(* Logix 5000 project; controller PLC_MCC1300_75F1 vendor 1 type 14 code 166 rev 32.11; software revision 32.04; part 5 of 83 *)
(* tags used below, declared in another part *)
   GP_PlateYPosition : GP_PlateYPosition;
   GP_PosWindow : GP_PosWindow;
   GP_RampManagement : GP_RampManagement;
   GP_RampSpace : GP_RampSpace;
   GP_ScadaPlate : GP_ScadaPlate;
   Gp_SpaceConvUtilities_V1 : GP_SpaceConvUtilities_V1;
   GP_TrackingAddCap : GP_TrackingAddCap;
   GP_TrackingFiring : GP_TrackingFiring;
   GP_TrackingFiringForConvoy : GP_TrackingFiringForConvoy;
   GP_TrackingGetFirstPlateInConveyor : GP_TrackingGetFirstPlateInConveyor;

ADD_ON_INSTRUCTION GP_PlateYPosition   (* revision 1.0 *)
VAR_IN_OUT
   INO_tPlateData : UDT_ConvoyCap_ZC; {required}
END_VAR
VAR_INPUT
   IN_dRequestGapLite_cmm : DINT; {access None, required}   // Requested gap between lites
   IN_dOffset_cmm : DINT; {access None, required}   // Position offset
   IN_xWander : BOOL; {access None, required}   // Calculate wander & total width
   IN_xBarycenter : BOOL; {access None, required}   // Calculate Barycenter
   IN_rgxNoGapLite : DINT; {access None, required}   // Consider gap of single lite [0:ConsiderGap, 1:NotConsiderGap]
END_VAR
VAR
   TMP_dLite : DINT; {access None}
   TMP_dMaxLites : DINT; {access None}
   TMP_dCapEdge_cmm : DINT; {access None}
END_VAR

ROUTINE Logic   (* structured text *)
   
   SIZE(INO_tPlateData.rgtCap[0].rgtLite[0],0,TMP_dMaxLites);
   IF INO_tPlateData.rgtCap[0].dID <> 0 THEN
       IF INO_tPlateData.rgtCap[0].dNumLites > 0 AND IN_xBarycenter THEN
           TMP_dCapEdge_cmm := (IN_dOffset_cmm + INO_tPlateData.rgtCap[0].dCutWander_cmm) - (INO_tPlateData.rgtCap[0].dWidth_cmm / 2) - (IN_dRequestGapLite_cmm / 2);
           FOR TMP_dLite := 0 TO TMP_dMaxLites - 1 DO
               IF INO_tPlateData.rgtCap[0].rgtLite[TMP_dLite].dID <> 0 THEN
                   INO_tPlateData.rgtCap[0].rgtLite[TMP_dLite].dBarycenter_cmm := TMP_dCapEdge_cmm + (INO_tPlateData.rgtCap[0].rgtLite[TMP_dLite].dWidth_cmm / 2);
                   IF NOT (IN_rgxNoGapLite.[TMP_dLite]) THEN
                       TMP_dCapEdge_cmm := TMP_dCapEdge_cmm + INO_tPlateData.rgtCap[0].rgtLite[TMP_dLite].dWidth_cmm + IN_dRequestGapLite_cmm;
   					//Update gap in cap data
   					INO_tPlateData.rgtCap[0].dGap_cmm := IN_dRequestGapLite_cmm;
                   ELSE
                       TMP_dCapEdge_cmm := TMP_dCapEdge_cmm + INO_tPlateData.rgtCap[0].rgtLite[TMP_dLite].dWidth_cmm;
                   END_IF;
               END_IF;
           END_FOR;
       ELSIF INO_tPlateData.rgtCap[0].dNumLites > 0 AND IN_xWander THEN
           FOR TMP_dLite := 0 TO TMP_dMaxLites - 1 DO
               IF INO_tPlateData.rgtCap[0].rgtLite[TMP_dLite].dID <> 0 THEN
                   TMP_dCapEdge_cmm := INO_tPlateData.rgtCap[0].rgtLite[TMP_dLite].dBarycenter_cmm - (INO_tPlateData.rgtCap[0].rgtLite[TMP_dLite].dWidth_cmm / 2);
               END_IF;
           END_FOR;
           FOR TMP_dLite := 0 TO TMP_dMaxLites - 1 DO
               IF INO_tPlateData.rgtCap[0].rgtLite[TMP_dLite].dID <> 0 THEN
                   INO_tPlateData.rgtCap[0].dWidth_cmm := (INO_tPlateData.rgtCap[0].rgtLite[TMP_dLite].dBarycenter_cmm + (INO_tPlateData.rgtCap[0].rgtLite[TMP_dLite].dWidth_cmm / 2)) - TMP_dCapEdge_cmm;
               END_IF;
           END_FOR;
           INO_tPlateData.rgtCap[0].dCutWander_cmm := (TMP_dCapEdge_cmm + (INO_tPlateData.rgtCap[0].dWidth_cmm / 2)) - IN_dOffset_cmm;
       END_IF;
   END_IF;
   
END_ROUTINE
END_ADD_ON_INSTRUCTION

ADD_ON_INSTRUCTION GP_PosWindow   (* revision 1.0 *)
VAR_INPUT
   IN_dTarget : DINT; {access None, required}   // Request position [user unit]
   IN_dActual : DINT; {access None, required}   // Actual position [user unit]
   IN_dTollerance : DINT; {access None, required}   // Tollerance window [user unit]
   IN_dMode : DINT; {access None, required}   // Type mode (0=Included, 1=Greater/Included, 2=Less/Includedl, 3=Greater, 4=Less)
END_VAR
VAR_OUTPUT
   OUT_xPositionReached : BOOL; {access None, required}   // Position reached
END_VAR
VAR
   TMP_dMaxValue : DINT; {access None}
   TMP_dMinValue : DINT; {access None}
END_VAR

ROUTINE Logic   (* structured text *)
   TMP_dMinValue := IN_dTarget - IN_dTollerance ;
   TMP_dMaxValue := IN_dTarget + IN_dTollerance ;
   
   CASE IN_dMode OF
   
   0:	IF IN_dActual >= TMP_dMinValue AND IN_dActual <= TMP_dMaxValue THEN
   
   		OUT_xPositionReached := 1 ;
   
   	ELSE
   
   		OUT_xPositionReached := 0 ;
   
   	END_IF;
   
   1:	IF IN_dActual >= TMP_dMinValue THEN
   
   		OUT_xPositionReached := 1 ;
   
   	ELSE
   
   		OUT_xPositionReached := 0 ;
   
   	END_IF;
   
   2:	IF IN_dActual <= TMP_dMaxValue THEN
   
   		OUT_xPositionReached := 1 ;
   
   	ELSE
   
   		OUT_xPositionReached := 0 ;
   
   	END_IF;
   
   3:	IF IN_dActual > TMP_dMinValue THEN
   
   		OUT_xPositionReached := 1 ;
   
   	ELSE
   
   		OUT_xPositionReached := 0 ;
   
   	END_IF;
   
   4:	IF IN_dActual < TMP_dMaxValue THEN
   
   		OUT_xPositionReached := 1 ;
   
   	ELSE
   
   		OUT_xPositionReached := 0 ;
   
   	END_IF;
   
   END_CASE;
   
   EnableOut := 1 ;
END_ROUTINE
END_ADD_ON_INSTRUCTION

ADD_ON_INSTRUCTION GP_RampManagement   (* revision 1.0 *)
VAR_INPUT
   IN_xRun : BOOL; {access None, required}   // Run command
   IN_dSpeed_Setpoint : DINT; {access None, required}   // Setpoint speed [mm/min]
   IN_rAcc : REAL; {access None, required}   // Acceleration [m/s2]
   IN_rDec : REAL; {access None, required}   // Deceleration [m/s2]
   IN_rScan : REAL; {access None, required}   // Previous scan [ms]
END_VAR
VAR_IN_OUT
   INO_rPV_Speed : REAL; {required}   // Processed speed value [mm/min]
END_VAR
VAR_OUTPUT
   OUT_dStep_cmm : DINT; {access None, required}   // Incremental step for each scan cycle [mm/100]
   OUT_xRampInProgress : BOOL; {access None, required}   // Acceleration/Deceleration ramp in progress
   OUT_xAccInProgress : BOOL; {access None, required}   // Acceleration ramp in progress
   OUT_xDecInProgress : BOOL; {access None, required}   // Deceleration ramp in progress
END_VAR
VAR_IN_OUT
   INO_rReminderStep : REAL; {required}   // Reminder Step [mm/min]
END_VAR
VAR
   TMP_rDecLim : REAL; {access None}   // Deceleration limit [mm/min]
   TMP_rAccLim : REAL; {access None}   // Acceleration limit [mm/min]
   TMP_rDecStep : REAL; {access None}   // Deceleration step [mm/min]
   TMP_rAccStep : REAL; {access None}   // Acceleration step [mm/min]
   TMP_rSpeed_Setpoint : REAL; {access None}   // Setpoint speed [mm/min]
   TMP_rScan : REAL; {access None}   // Previous scan [ms]
   TMP_rStep : REAL; {access None}   // Actual Step with reminder [mm/min]
   TMP_rStepRound : REAL; {access None}   // Actual Step with reminder [mm/min]
END_VAR

ROUTINE Logic   (* structured text *)
   //Initialize
   OUT_dStep_cmm := 0;
   TMP_rSpeed_Setpoint := IN_dSpeed_Setpoint;
   TMP_rScan := IN_rScan;
   OUT_xRampInProgress := 0;
   OUT_xAccInProgress := 0;
   OUT_xDecInProgress := 0;
   
   //Check Speed, Acceleration and Deceleration Values > 0
   
   IF TMP_rSpeed_Setpoint > 0.0 AND IN_rAcc > 0.0 AND IN_rDec > 0.0 THEN
   
       // Acceleration
       IF IN_xRun AND TMP_rSpeed_Setpoint > INO_rPV_Speed THEN
           TMP_rAccStep := IN_rAcc * TMP_rScan * 60.0;
           INO_rPV_Speed := INO_rPV_Speed + TMP_rAccStep;
           TMP_rAccLim := TMP_rSpeed_Setpoint + TMP_rAccStep;
           OUT_xRampInProgress := 1;
           OUT_xAccInProgress := 1;
   
           IF IN_xRun AND INO_rPV_Speed > TMP_rSpeed_Setpoint AND INO_rPV_Speed < TMP_rAccLim THEN
               INO_rPV_Speed := TMP_rSpeed_Setpoint;
           END_IF;
   
           // Deceleration
   
       ELSIF (IN_xRun AND TMP_rSpeed_Setpoint < INO_rPV_Speed) OR (NOT (IN_xRun) AND INO_rPV_Speed > 0.0) THEN
           TMP_rDecStep := IN_rDec * TMP_rScan * 60.0;
           INO_rPV_Speed := INO_rPV_Speed - TMP_rDecStep;
           TMP_rDecLim := TMP_rSpeed_Setpoint - TMP_rDecStep;
           OUT_xRampInProgress := 1;
           OUT_xDecInProgress := 1;
   
           IF IN_xRun AND INO_rPV_Speed < TMP_rSpeed_Setpoint AND INO_rPV_Speed > TMP_rDecLim THEN
               INO_rPV_Speed := TMP_rSpeed_Setpoint;
           END_IF;
       END_IF;
   
       // Delete PV_Speed If < 0
   
       IF INO_rPV_Speed < 0.0 THEN
           INO_rPV_Speed := 0.0;
       END_IF;
   
   	// Calculate step value
   	TMP_rStep := ((INO_rPV_Speed * TMP_rScan) / 600.0) + INO_rReminderStep;
   
   	// Calculate the round value
   	TMP_rStepRound := TRUNC(TMP_rStep + 0.5);
   	OUT_dStep_cmm := TRUNC(TMP_rStep + 0.5);
   
       // Save the reminder for the next cycle
       INO_rReminderStep := TMP_rStep - TMP_rStepRound;
   
   END_IF;
END_ROUTINE
END_ADD_ON_INSTRUCTION

ADD_ON_INSTRUCTION GP_RampSpace   (* revision 1.0 *)
VAR_INPUT
   IN_rAcc_m_s2 : REAL; {access None, required}   // Acceleration ramp [m/s2]
   IN_rDec_m_s2 : REAL; {access None, required}   // Deceleration ramp [m/s2]
   IN_dActualSpeed_mm_min : DINT; {access None, required}   // Actual speed [mm/min]
END_VAR
VAR_OUTPUT
   OUT_dAccSpace_cmm : DINT; {access None, required}   // Acceleration space [mm/100]
   OUT_dDecSpace_cmm : DINT; {access None, required}   // Deceleration space [mm/100]
END_VAR
VAR
   TMP_rDec_mm_s2 : REAL; {access None}   // Deceleration ramp [mm/s2]
   TMP_rAcc_mm_s2 : REAL; {access None}   // Acceleration ramp [mm/s2]
   TMP_dAcc_mm_s2 : DINT; {access None}   // Acceleration ramp [mm/s2]
   TMP_dDec_mm_s2 : DINT; {access None}   // Deceleration ramp [mm/s2]
END_VAR

ROUTINE Logic   (* structured text *)
   //Calculate Acceleration and deceleration space
   
   //Acceleration
   TMP_rAcc_mm_s2 := IN_rAcc_m_s2 * 1000.0;
   TMP_dAcc_mm_s2 := TMP_rAcc_mm_s2;
   //Deceleration
   TMP_rDec_mm_s2 := IN_rDec_m_s2 * 1000.0;
   TMP_dDec_mm_s2 := TMP_rDec_mm_s2;
   
   OUT_dAccSpace_cmm:= (((IN_dActualSpeed_mm_min / 60)*(IN_dActualSpeed_mm_min / 60))/(2*TMP_dAcc_mm_s2)) * 100;
   OUT_dDecSpace_cmm:= (((IN_dActualSpeed_mm_min / 60)*(IN_dActualSpeed_mm_min / 60))/(2*TMP_dDec_mm_s2)) * 100;
END_ROUTINE
END_ADD_ON_INSTRUCTION

ADD_ON_INSTRUCTION GP_Rotator   (* revision 1.0 *)
VAR_IN_OUT
   STC_tLogics : MAC_Rotator; {required}   // Logics Tags
        .PH_x.0   // Rise frame
        .PH_x.3   // End rise
        .PH_x.11   // End rotation Cw
        .PH_x.12   // Rotation counterclockwise
        .PH_x.15   // End rotation Ccw
        .PH_x.4   // Descent frame
        .PH_x.7   // End descent
        .PH_x.8   // Rotation clockwise
   STC_tHMR : MAC_Rotator_HMR; {required}   // HMI Tags
        .rgxMan.0   // Rise
        .rgxMan.1   // Descent
        .rgxMan.10   // Clockwise rotation jog
        .rgxMan.11   // Counter Clockwise rotation jog
        .rgxMan.14   // Enable brake release
        .rgxMan.15   // Disable brake release
        .rgxMan.8   // Clockwise rotation
        .rgxMan.9   // Counter Clockwise rotation
   STC_tHMW : MAC_Rotator_HMW; {required}   // HMI Tags
        .rgxMan.0   // Rise
        .rgxMan.1   // Descent
        .rgxMan.10   // Clockwise rotation jog
        .rgxMan.11   // Counter Clockwise rotation jog
        .rgxMan.14   // Enable brake release
        .rgxMan.15   // Disable brake release
        .rgxMan.8   // Clockwise rotation
        .rgxMan.9   // Counter Clockwise rotation
   STC_tData : UDT_Convoy_SL; {required}   // Plate data
END_VAR
VAR_INPUT
   IN_xCycleON : BOOL; {access None, required}   // Zone cycle ON
   IN_xPhaseAdvancement : BOOL; {access None, required}   // Condition OK for phases advancement
   IN_xManualMode : BOOL; {access None, required}   // Manual mode enabled
   IN_xReqAccess : BOOL; {access None}   // Request access area
   IN_xDoneAccess : BOOL; {access None}   // Done access area
   IN_iOpSide : INT; {access None, visible}   // Operator side (0=Right side 1=Left side)
   IN_dWander_cmm : DINT; {access None}   // Convoy wander [mm/100] (Optional 0 = No wander)
   IN_xConditionToDescent : BOOL; {access None}
   IN_xDriveFeedback : BOOL; {access None}
   IN_xHighPosition : BOOL; {access None}
   IN_xLowPosition : BOOL; {access None}
   IN_xPositionReached : BOOL; {access None}
   IN_dRotatorPosition_cdeg : DINT; {access None}
END_VAR
VAR_IN_OUT
   INO_tFlags : WorkingFlags_Rotator; {required}
   INO_dPlatePosition_cmm : DINT; {required}   // Plate position [mm/100]
END_VAR
VAR_INPUT
   OUT_xDriveEnable : BOOL; {access None}   // (Only for HMRm)
   OUT_xRun : BOOL; {access None}   // (Only for HMRm)
   OUT_xReverse : BOOL; {access None}   // (Only for HMRm)
   OUT_xRise : BOOL; {access None}   // (Only for HMRm)
   OUT_xDescent : BOOL; {access None}   // (Only for HMRm)
   OUT_xBrakeRelease : BOOL; {access None}   // (Only for HMRm)
END_VAR
VAR
   TMP_rWeight_kg : REAL; {access None}
   TMP_iPointerLite : INT; {access None}
   TMP_iSizeCap : INT; {access None}
   TMP_iPointerCap : INT; {access None}
   TMP_iSizeLite : INT; {access None}
   TMP_iStepNumber : INT; {access None}   // Step number of rotation
   TMP_dEdgeToCenter_cmm : DINT; {access None}   // Distance between convoy edge and center rotator [mm/100]
END_VAR

ROUTINE Logic   (* ladder *)
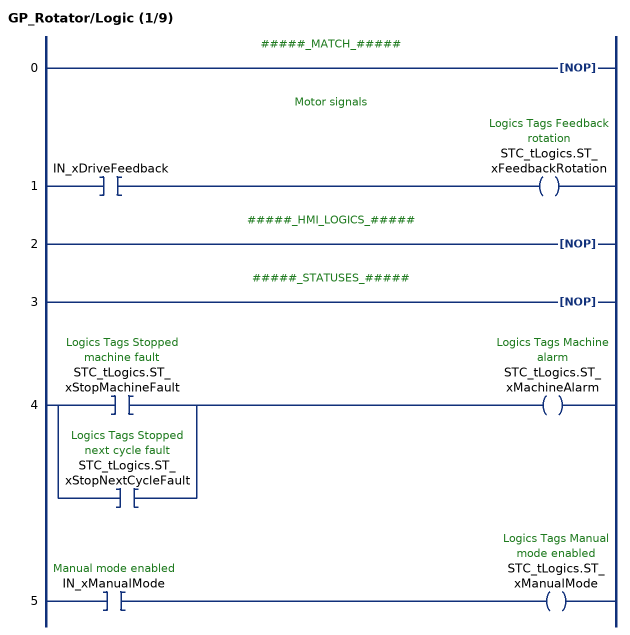
   // #####_MATCH_#####
   0: NOP();
   // Motor signals
   1: XIC(IN_xDriveFeedback)OTE(STC_tLogics.ST_xFeedbackRotation);
   // #####_HMI_LOGICS_#####
   2: NOP();
   // #####_STATUSES_#####
   3: NOP();
   4: [XIC(STC_tLogics.ST_xStopMachineFault) ,XIC(STC_tLogics.ST_xStopNextCycleFault) ]OTE(STC_tLogics.ST_xMachineAlarm);
   5: XIC(IN_xManualMode)OTE(STC_tLogics.ST_xManualMode);
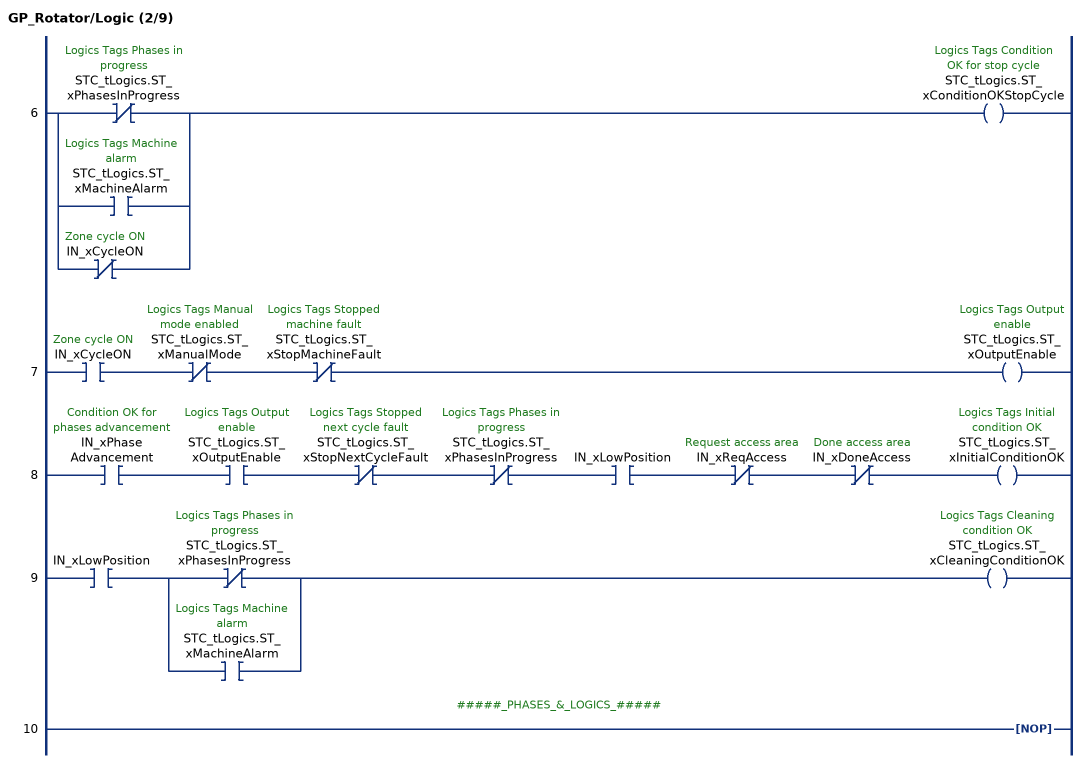
   6: [XIO(STC_tLogics.ST_xPhasesInProgress) ,XIC(STC_tLogics.ST_xMachineAlarm) ,XIO(IN_xCycleON) ]OTE(STC_tLogics.ST_xConditionOKStopCycle);
   7: XIC(IN_xCycleON)XIO(STC_tLogics.ST_xManualMode)XIO(STC_tLogics.ST_xStopMachineFault)OTE(STC_tLogics.ST_xOutputEnable);
   8: XIC(IN_xPhaseAdvancement)XIC(STC_tLogics.ST_xOutputEnable)XIO(STC_tLogics.ST_xStopNextCycleFault)XIO(STC_tLogics.ST_xPhasesInProgress)XIC(IN_xLowPosition)XIO(IN_xReqAccess)XIO(IN_xDoneAccess)OTE(STC_tLogics.ST_xInitialConditionOK);
   9: XIC(IN_xLowPosition)[XIO(STC_tLogics.ST_xPhasesInProgress) ,XIC(STC_tLogics.ST_xMachineAlarm) ]OTE(STC_tLogics.ST_xCleaningConditionOK);
   // #####_PHASES_&_LOGICS_#####
   10: NOP();
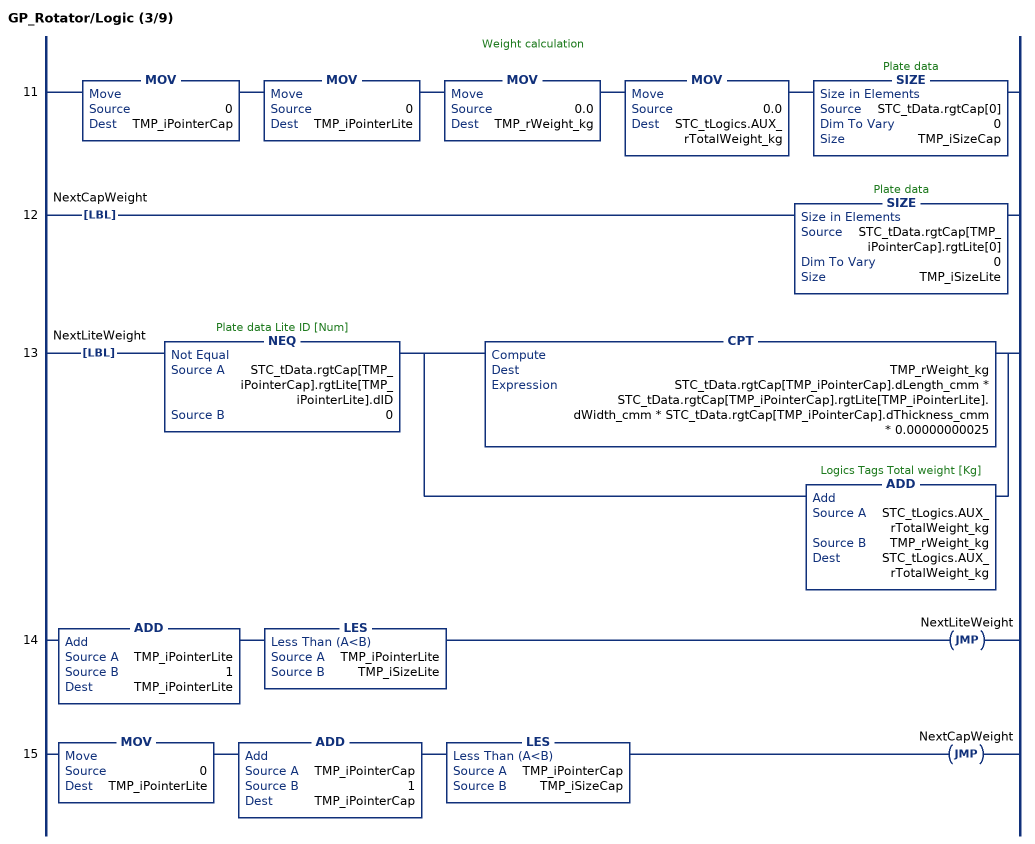
   // Weight calculation
   11: MOV(0,TMP_iPointerCap)MOV(0,TMP_iPointerLite)MOV(0.0,TMP_rWeight_kg)MOV(0.0,STC_tLogics.AUX_rTotalWeight_kg)SIZE(STC_tData.rgtCap[0],0,TMP_iSizeCap);
   12: LBL(NextCapWeight)SIZE(STC_tData.rgtCap[TMP_iPointerCap].rgtLite[0],0,TMP_iSizeLite);
   13: LBL(NextLiteWeight)NEQ(STC_tData.rgtCap[TMP_iPointerCap].rgtLite[TMP_iPointerLite].dID,0)[CPT(TMP_rWeight_kg,STC_tData.rgtCap[TMP_iPointerCap].dLength_cmm * STC_tData.rgtCap[TMP_iPointerCap].rgtLite[TMP_iPointerLite].dWidth_cmm * STC_tData.rgtCap[TMP_iPointerCap].dThickness_cmm * 0.00000000025) ,ADD(STC_tLogics.AUX_rTotalWeight_kg,TMP_rWeight_kg,STC_tLogics.AUX_rTotalWeight_kg) ];
   14: ADD(TMP_iPointerLite,1,TMP_iPointerLite)LES(TMP_iPointerLite,TMP_iSizeLite)JMP(NextLiteWeight);
   15: MOV(0,TMP_iPointerLite)ADD(TMP_iPointerCap,1,TMP_iPointerCap)LES(TMP_iPointerCap,TMP_iSizeCap)JMP(NextCapWeight);
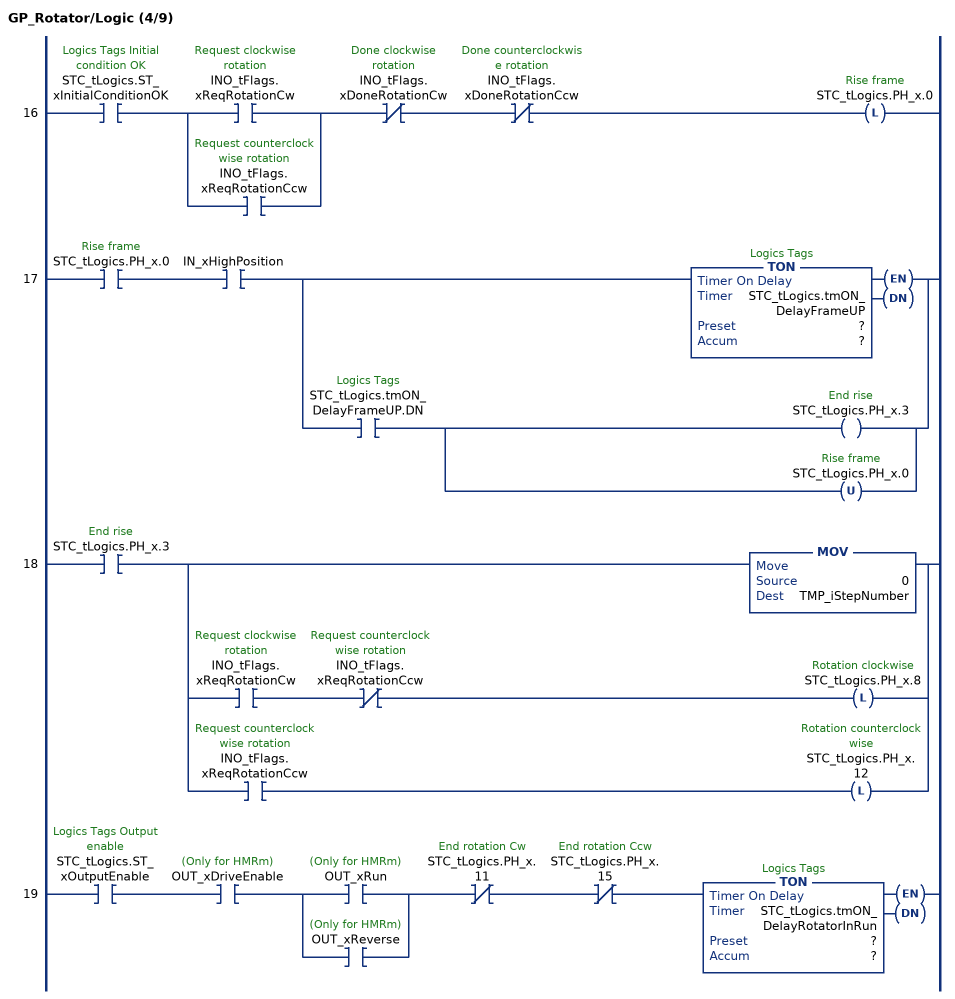
   16: XIC(STC_tLogics.ST_xInitialConditionOK)[XIC(INO_tFlags.xReqRotationCw) ,XIC(INO_tFlags.xReqRotationCcw) ]XIO(INO_tFlags.xDoneRotationCw)XIO(INO_tFlags.xDoneRotationCcw)OTL(STC_tLogics.PH_x.0);
   17: XIC(STC_tLogics.PH_x.0)XIC(IN_xHighPosition)[TON(STC_tLogics.tmON_DelayFrameUP,?,?) ,XIC(STC_tLogics.tmON_DelayFrameUP.DN) [OTE(STC_tLogics.PH_x.3) ,OTU(STC_tLogics.PH_x.0) ] ];
   18: XIC(STC_tLogics.PH_x.3)[MOV(0,TMP_iStepNumber) ,XIC(INO_tFlags.xReqRotationCw) XIO(INO_tFlags.xReqRotationCcw) OTL(STC_tLogics.PH_x.8) ,XIC(INO_tFlags.xReqRotationCcw) OTL(STC_tLogics.PH_x.12) ];
   19: XIC(STC_tLogics.ST_xOutputEnable)XIC(OUT_xDriveEnable)[XIC(OUT_xRun) ,XIC(OUT_xReverse) ]XIO(STC_tLogics.PH_x.11)XIO(STC_tLogics.PH_x.15)TON(STC_tLogics.tmON_DelayRotatorInRun,?,?);
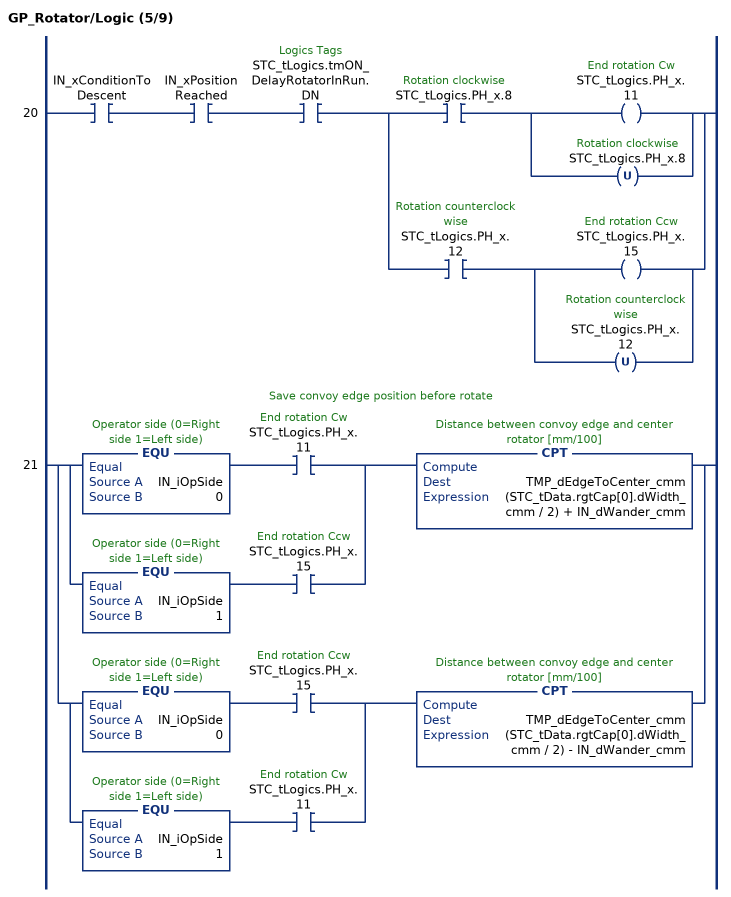
   20: XIC(IN_xConditionToDescent)XIC(IN_xPositionReached)XIC(STC_tLogics.tmON_DelayRotatorInRun.DN)[XIC(STC_tLogics.PH_x.8) [OTE(STC_tLogics.PH_x.11) ,OTU(STC_tLogics.PH_x.8) ] ,XIC(STC_tLogics.PH_x.12) [OTE(STC_tLogics.PH_x.15) ,OTU(STC_tLogics.PH_x.12) ] ];
   // Save convoy edge position before rotate
   21: [[EQU(IN_iOpSide,0) XIC(STC_tLogics.PH_x.11) ,EQU(IN_iOpSide,1) XIC(STC_tLogics.PH_x.15) ] CPT(TMP_dEdgeToCenter_cmm,(STC_tData.rgtCap[0].dWidth_cmm / 2) + IN_dWander_cmm) ,[EQU(IN_iOpSide,0) XIC(STC_tLogics.PH_x.15) ,EQU(IN_iOpSide,1) XIC(STC_tLogics.PH_x.11) ] CPT(TMP_dEdgeToCenter_cmm,(STC_tData.rgtCap[0].dWidth_cmm / 2) - IN_dWander_cmm) ];
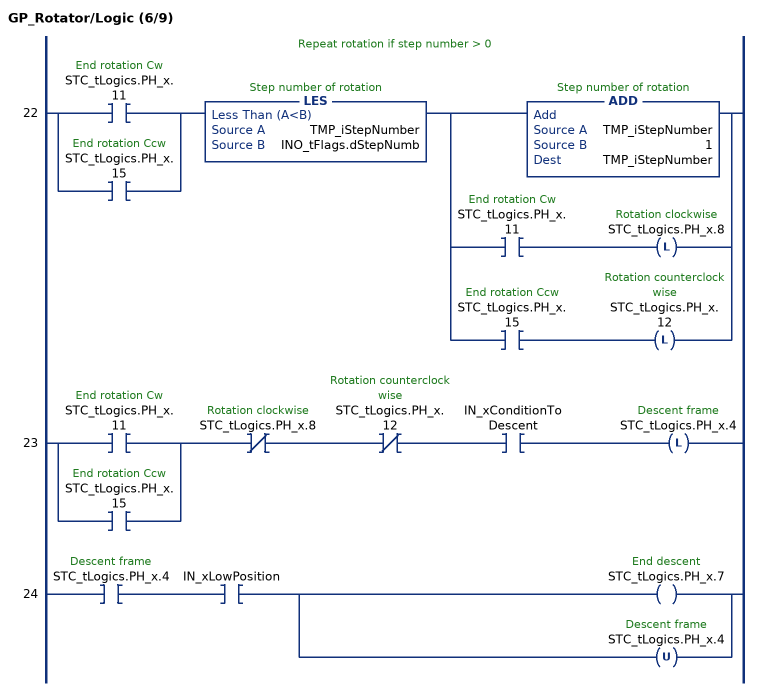
   // Repeat rotation if step number > 0
   22: [XIC(STC_tLogics.PH_x.11) ,XIC(STC_tLogics.PH_x.15) ]LES(TMP_iStepNumber,INO_tFlags.dStepNumb)[ADD(TMP_iStepNumber,1,TMP_iStepNumber) ,XIC(STC_tLogics.PH_x.11) OTL(STC_tLogics.PH_x.8) ,XIC(STC_tLogics.PH_x.15) OTL(STC_tLogics.PH_x.12) ];
   23: [XIC(STC_tLogics.PH_x.11) ,XIC(STC_tLogics.PH_x.15) ]XIO(STC_tLogics.PH_x.8)XIO(STC_tLogics.PH_x.12)XIC(IN_xConditionToDescent)OTL(STC_tLogics.PH_x.4);
   24: XIC(STC_tLogics.PH_x.4)XIC(IN_xLowPosition)[OTE(STC_tLogics.PH_x.7) ,OTU(STC_tLogics.PH_x.4) ];
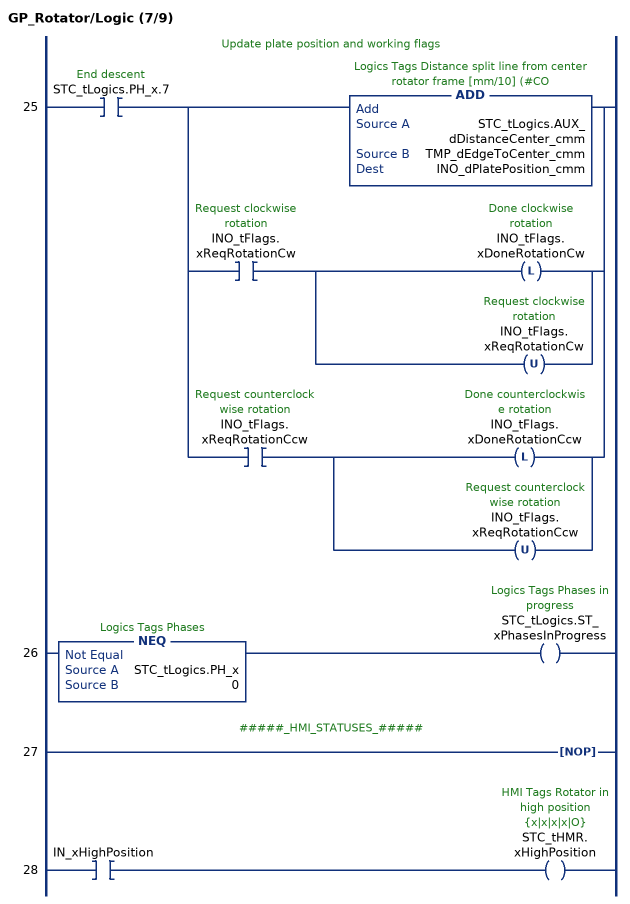
   // Update plate position and working flags
   25: XIC(STC_tLogics.PH_x.7)[ADD(STC_tLogics.AUX_dDistanceCenter_cmm,TMP_dEdgeToCenter_cmm,INO_dPlatePosition_cmm) ,XIC(INO_tFlags.xReqRotationCw) [OTL(INO_tFlags.xDoneRotationCw) ,OTU(INO_tFlags.xReqRotationCw) ] ,XIC(INO_tFlags.xReqRotationCcw) [OTL(INO_tFlags.xDoneRotationCcw) ,OTU(INO_tFlags.xReqRotationCcw) ] ];
   26: NEQ(STC_tLogics.PH_x,0)OTE(STC_tLogics.ST_xPhasesInProgress);
   // #####_HMI_STATUSES_#####
   27: NOP();
   28: XIC(IN_xHighPosition)OTE(STC_tHMR.xHighPosition);
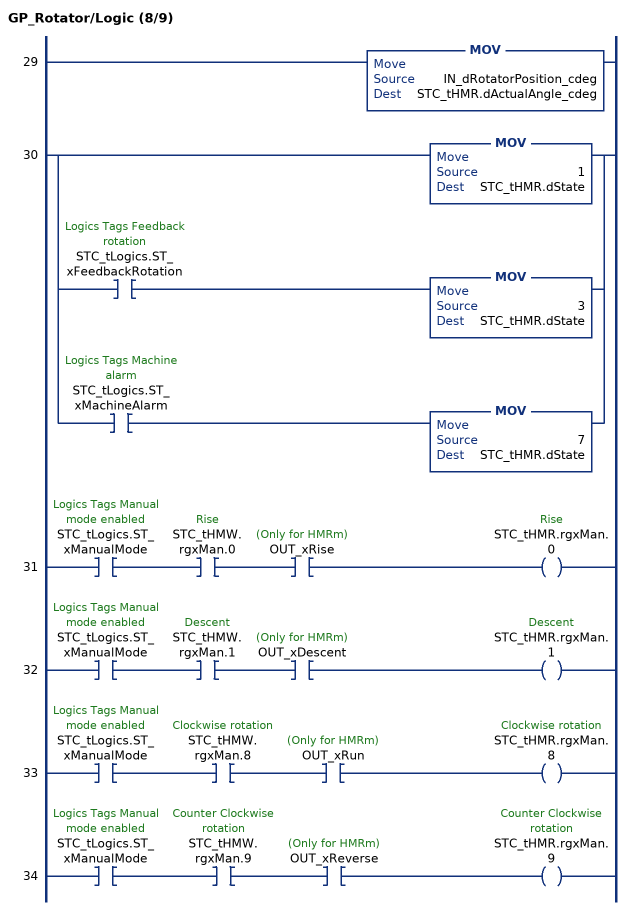
   29: MOV(IN_dRotatorPosition_cdeg,STC_tHMR.dActualAngle_cdeg);
   30: [MOV(1,STC_tHMR.dState) ,XIC(STC_tLogics.ST_xFeedbackRotation) MOV(3,STC_tHMR.dState) ,XIC(STC_tLogics.ST_xMachineAlarm) MOV(7,STC_tHMR.dState) ];
   31: XIC(STC_tLogics.ST_xManualMode)XIC(STC_tHMW.rgxMan.0)XIC(OUT_xRise)OTE(STC_tHMR.rgxMan.0);
   32: XIC(STC_tLogics.ST_xManualMode)XIC(STC_tHMW.rgxMan.1)XIC(OUT_xDescent)OTE(STC_tHMR.rgxMan.1);
   33: XIC(STC_tLogics.ST_xManualMode)XIC(STC_tHMW.rgxMan.8)XIC(OUT_xRun)OTE(STC_tHMR.rgxMan.8);
   34: XIC(STC_tLogics.ST_xManualMode)XIC(STC_tHMW.rgxMan.9)XIC(OUT_xReverse)OTE(STC_tHMR.rgxMan.9);
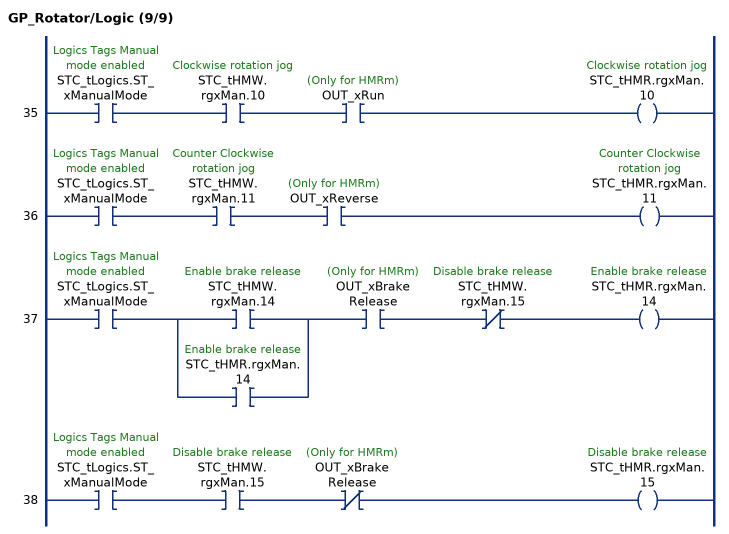
   35: XIC(STC_tLogics.ST_xManualMode)XIC(STC_tHMW.rgxMan.10)XIC(OUT_xRun)OTE(STC_tHMR.rgxMan.10);
   36: XIC(STC_tLogics.ST_xManualMode)XIC(STC_tHMW.rgxMan.11)XIC(OUT_xReverse)OTE(STC_tHMR.rgxMan.11);
   37: XIC(STC_tLogics.ST_xManualMode)[XIC(STC_tHMW.rgxMan.14) ,XIC(STC_tHMR.rgxMan.14) ]XIC(OUT_xBrakeRelease)XIO(STC_tHMW.rgxMan.15)OTE(STC_tHMR.rgxMan.14);
   38: XIC(STC_tLogics.ST_xManualMode)XIC(STC_tHMW.rgxMan.15)XIO(OUT_xBrakeRelease)OTE(STC_tHMR.rgxMan.15);
END_ROUTINE
END_ADD_ON_INSTRUCTION

ADD_ON_INSTRUCTION GP_ScadaPlate   (* revision 1.0 *)
VAR_IN_OUT
   IN_tPlate : UDT_Convoy_SL; {required}
END_VAR
VAR_INPUT
   IN_iIndexArray : DINT; {required}
   IN_dHeadPosition_cmm : DINT; {required}
   IN_dConveyorWidht_cmm : DINT; {required}
   IN_dConveyorLenght_cmm : DINT; {required}
   IN_xLastModalityLoadBkw : BOOL; {required}
   IN_xLastModalityUnloadBkw : BOOL; {required}
   IN_xYWithBaricentre : BOOL; {required}
   IN_xYInversionLite : BOOL; {required}   // AtoX
END_VAR
VAR_IN_OUT
   Scada_Plate : HMI_LiteData[5,2,7]; {required}
END_VAR
VAR_OUTPUT
   DebugOut : DINT; {access None}
END_VAR
VAR
   TMP_dCapClean : DINT; {access None}
   TMP_dLiteClean : DINT; {access None}
   TMP_dWidth_mm : DINT; {access None}
   TMP_dLiteInv : DINT; {access None}
   TMP_dConveyorLenght : DINT; {access None}
   TMP_dCountDest : DINT; {access None}
   TMP_dMaxLite : DINT; {access None}
   TMP_dMaxCap : DINT; {access None}
   TMP_dHeadPosition_mm : DINT; {access None}
   TMP_dLite : DINT; {access None}
   TMP_dCap : DINT; {access None}
   Debug : DINT[32]; {access None}
END_VAR

ROUTINE Logic   (* structured text *)
   //////////////////////////////////////////////////////////
   //   Copyright (c)  <Key Automation srl>
   //------------------------------------------------------------
   //   Routine: <Routine Name>
   //   Author: <Developer Name>
   //   Created: <Date>
   //------------------------------------------------------------
   //   Description:
   //           <Description>
   
   //   History:
   
   ////////////////////////////////////////////////////////////
   
   //Size arrays
   
   size(IN_tPlate.rgtCap,0,TMP_dMaxCap);
   size(IN_tPlate.rgtCap[0].rgtLite,0,TMP_dMaxLite);
   
   //Cleaning Data
   
   FOR TMP_dCap := 0 TO TMP_dMaxCap - 1 DO
       FOR TMP_dLite := 0 TO TMP_dMaxLite - 1 DO
   		Scada_Plate[IN_iIndexArray, TMP_dCap, TMP_dLite].dTail_PosX_mm := 0;
   		Scada_Plate[IN_iIndexArray, TMP_dCap, TMP_dLite].dPlateLength_mm := 0;
   		Scada_Plate[IN_iIndexArray, TMP_dCap, TMP_dLite].dPositionY_mm := 0;
   		Scada_Plate[IN_iIndexArray, TMP_dCap, TMP_dLite].dPlateWidth_mm := 0;
   		Scada_Plate[IN_iIndexArray, TMP_dCap, TMP_dLite].dDestination := 0;
   		Scada_Plate[IN_iIndexArray, TMP_dCap, TMP_dLite].dAlternative := 0;
   		Scada_Plate[IN_iIndexArray, TMP_dCap, TMP_dLite].dSecondDestination := 0;
   		Scada_Plate[IN_iIndexArray, TMP_dCap, TMP_dLite].dPlateId := 0;
   		Scada_Plate[IN_iIndexArray, TMP_dCap, TMP_dLite].dProductionID := 0;
       END_FOR;
   END_FOR;
   
   //Write data
   //Calculate Head Position
   TMP_dHeadPosition_mm := IN_dHeadPosition_cmm / 100;
   TMP_dConveyorLenght := IN_dConveyorLenght_cmm / 100;
   TMP_dWidth_mm := IN_dConveyorWidht_cmm / 100;
   
   FOR TMP_dCap := 0 TO TMP_dMaxCap - 1 DO
   	FOR TMP_dLite := 0 TO TMP_dMaxLite - 1 DO
   		IF IN_tPlate.rgtCap[TMP_dCap].rgtLite[TMP_dLite].dID <> 0 THEN
   			//Plate ID
   			Scada_Plate[IN_iIndexArray, TMP_dCap, TMP_dLite].dPlateId := IN_tPlate.rgtCap[TMP_dCap].rgtLite[TMP_dLite].dID;
   			//Production ID
   			Scada_Plate[IN_iIndexArray, TMP_dCap, TMP_dLite].dProductionID := IN_tPlate.rgtCap[TMP_dCap].rgtLite[TMP_dLite].dProductionID;
   			//Plate lenght
   			Scada_Plate[IN_iIndexArray, TMP_dCap, TMP_dLite].dPlateLength_mm := IN_tPlate.rgtCap[TMP_dCap].dLength_cmm / 100;
   			//Plate widht
   			Scada_Plate[IN_iIndexArray, TMP_dCap, TMP_dLite].dPlateWidth_mm := IN_tPlate.rgtCap[TMP_dCap].rgtLite[TMP_dLite].dWidth_cmm / 100;
   			//Destination
   			FOR TMP_dCountDest := 0 TO 32-1 DO
   				//Main Destination
   				IF IN_tPlate.rgtCap[TMP_dCap].rgtLite[TMP_dLite].tDestination.rgxMain.[TMP_dCountDest] THEN
   					Scada_Plate[IN_iIndexArray, TMP_dCap, TMP_dLite].dDestination := TMP_dCountDest+1;
   				END_IF;
   				//Source
   				//IF IN_tPlate.rgtCap[TMP_dCap].rgtLites[TMP_dLite].rgxOrigin[TMP_dCountDest] THEN
   				//    Scada_Plate[IN_iIndexArray, TMP_dCap, TMP_dLite].dSource := TMP_dCountDest;
   				//END_IF;
   				//Alternative Destination
   				IF IN_tPlate.rgtCap[TMP_dCap].rgtLite[TMP_dLite].tDestination.rgxAlternative.[TMP_dCountDest] THEN
   					Scada_Plate[IN_iIndexArray, TMP_dCap, TMP_dLite].dAlternative := TMP_dCountDest+1;
   				END_IF;
   				//Second Destination
   				IF IN_tPlate.rgtCap[TMP_dCap].rgtLite[TMP_dLite].tDestination.rgxSecChoice.[TMP_dCountDest] THEN
   					Scada_Plate[IN_iIndexArray, TMP_dCap, TMP_dLite].dSecondDestination := TMP_dCountDest+1;
   	 			END_IF;
   			END_FOR;
   			//IF IN_tPlate.rgtCap[TMP_dCap].rgtLites[TMP_dLite].tDestination.rgxMain[25] THEN //cullet
   			//	Scada_Plate[IN_iIndexArray, TMP_dCap, TMP_dLite].dDestination := 25;
   			//END_IF;
   			//Set origin to 0 in case of destination is <> 0
    			// IF Scada_Plate[IN_iIndexArray, TMP_dCap, TMP_dLite].dDestination <> 0 THEN
    			//	Scada_Plate[IN_iIndexArray, TMP_dCap, TMP_dLite].dSource := 0;
    			//END_IF;